(* Logix 5000 project; controller FV vendor 1 type 14 code 217 rev 31.11; software revision 31.00; part 21 of 63 *)
(* tags used below, declared in another part *)
   CheckTimeMask : INT;
   Delphi_Does_Eng_Func : BOOL;
   FR_FV28_AV01 : PlantItem;   // FV28_AV01
   FR_FV28_AV04 : PlantItem;   // FV28_AV04
   FR_FV28_AV05 : PlantItem;   // FV28_AV05
   FR_FV28_AV06 : PlantItem;   // FV28_AV06
   FR_FV28_AV07 : PlantItem;   // FV28_AV07
   FR_FV29_AV01 : PlantItem;   // FV29_AV01
   FR_FV29_AV04 : PlantItem;   // FV29_AV04
   FR_N255 : INT[265];   // CHECKWORDS
   FR_VB1_AV04 : PlantItem;   // VB1_AV04
   FR_VB1_AV05 : PlantItem;   // VB1_AV05
   FR_VB1_AV06 : PlantItem;   // VB1_AV06
   FR_VB1_AV07 : PlantItem;   // VB1_AV07
   FR_VB1_AV08 : PlantItem;   // VB1_AV08
   FR_VB1_AV09 : PlantItem;   // VB1_AV09
   TempChecktime : DINT;
(* FR_Common, continued *)

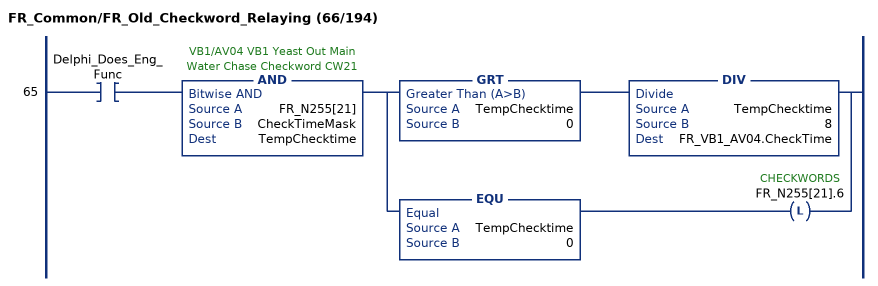
   [picture p370: FR_Common/FR_Old_Checkword_Relaying rungs 65-65]
   65: XIC(Delphi_Does_Eng_Func)AND(FR_N255[21],CheckTimeMask,TempChecktime)[GRT(TempChecktime,0) DIV(TempChecktime,8,FR_VB1_AV04.CheckTime) ,EQU(TempChecktime,0) OTL(FR_N255[21].6) ];
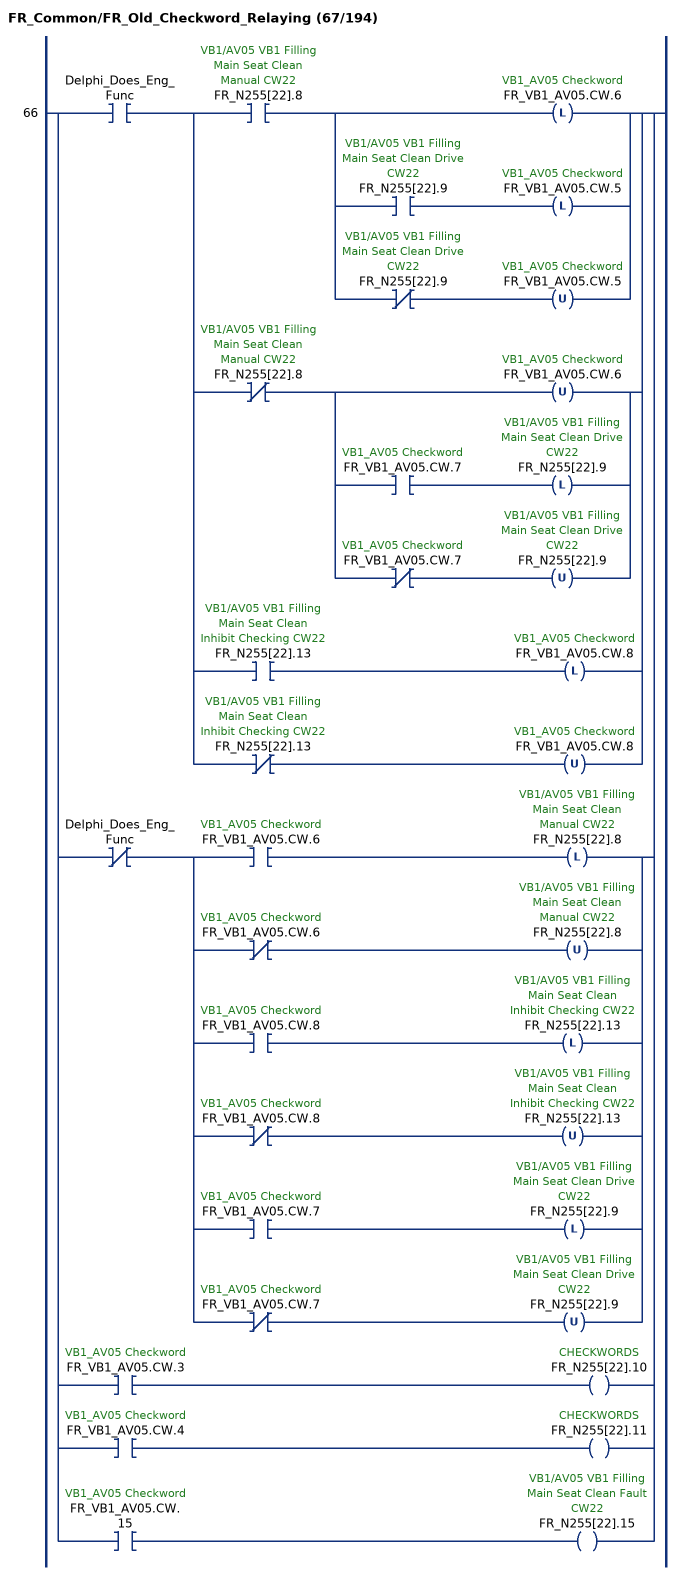
   66: [XIC(Delphi_Does_Eng_Func) [[XIC(FR_N255[22].8) [OTL(FR_VB1_AV05.CW.6) ,XIC(FR_N255[22].9) OTL(FR_VB1_AV05.CW.5) ,XIO(FR_N255[22].9) OTU(FR_VB1_AV05.CW.5) ] ,XIO(FR_N255[22].8) [OTU(FR_VB1_AV05.CW.6) ,[XIC(FR_VB1_AV05.CW.7) OTL(FR_N255[22].9) ,XIO(FR_VB1_AV05.CW.7) OTU(FR_N255[22].9) ] ] ] ,[XIC(FR_N255[22].13) OTL(FR_VB1_AV05.CW.8) ,XIO(FR_N255[22].13) OTU(FR_VB1_AV05.CW.8) ] ] ,XIO(Delphi_Does_Eng_Func) [[XIC(FR_VB1_AV05.CW.6) OTL(FR_N255[22].8) ,XIO(FR_VB1_AV05.CW.6) OTU(FR_N255[22].8) ] ,[XIC(FR_VB1_AV05.CW.8) OTL(FR_N255[22].13) ,XIO(FR_VB1_AV05.CW.8) OTU(FR_N255[22].13) ] ,[XIC(FR_VB1_AV05.CW.7) OTL(FR_N255[22].9) ,XIO(FR_VB1_AV05.CW.7) OTU(FR_N255[22].9) ] ] ,XIC(FR_VB1_AV05.CW.3) OTE(FR_N255[22].10) ,XIC(FR_VB1_AV05.CW.4) OTE(FR_N255[22].11) ,XIC(FR_VB1_AV05.CW.15) OTE(FR_N255[22].15) ];
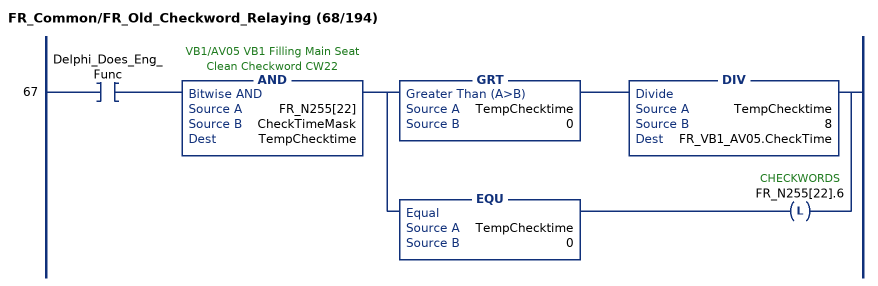
   67: XIC(Delphi_Does_Eng_Func)AND(FR_N255[22],CheckTimeMask,TempChecktime)[GRT(TempChecktime,0) DIV(TempChecktime,8,FR_VB1_AV05.CheckTime) ,EQU(TempChecktime,0) OTL(FR_N255[22].6) ];
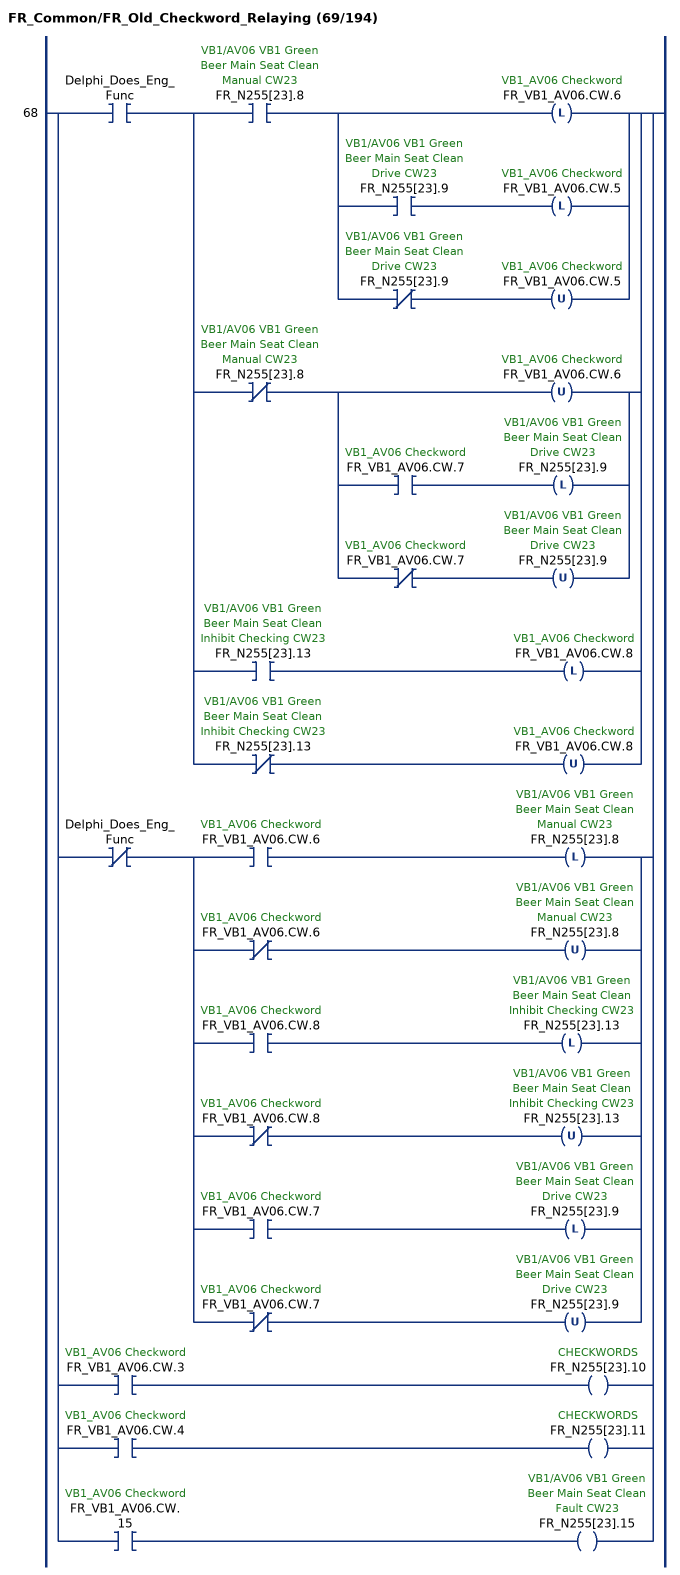
   68: [XIC(Delphi_Does_Eng_Func) [[XIC(FR_N255[23].8) [OTL(FR_VB1_AV06.CW.6) ,XIC(FR_N255[23].9) OTL(FR_VB1_AV06.CW.5) ,XIO(FR_N255[23].9) OTU(FR_VB1_AV06.CW.5) ] ,XIO(FR_N255[23].8) [OTU(FR_VB1_AV06.CW.6) ,[XIC(FR_VB1_AV06.CW.7) OTL(FR_N255[23].9) ,XIO(FR_VB1_AV06.CW.7) OTU(FR_N255[23].9) ] ] ] ,[XIC(FR_N255[23].13) OTL(FR_VB1_AV06.CW.8) ,XIO(FR_N255[23].13) OTU(FR_VB1_AV06.CW.8) ] ] ,XIO(Delphi_Does_Eng_Func) [[XIC(FR_VB1_AV06.CW.6) OTL(FR_N255[23].8) ,XIO(FR_VB1_AV06.CW.6) OTU(FR_N255[23].8) ] ,[XIC(FR_VB1_AV06.CW.8) OTL(FR_N255[23].13) ,XIO(FR_VB1_AV06.CW.8) OTU(FR_N255[23].13) ] ,[XIC(FR_VB1_AV06.CW.7) OTL(FR_N255[23].9) ,XIO(FR_VB1_AV06.CW.7) OTU(FR_N255[23].9) ] ] ,XIC(FR_VB1_AV06.CW.3) OTE(FR_N255[23].10) ,XIC(FR_VB1_AV06.CW.4) OTE(FR_N255[23].11) ,XIC(FR_VB1_AV06.CW.15) OTE(FR_N255[23].15) ];
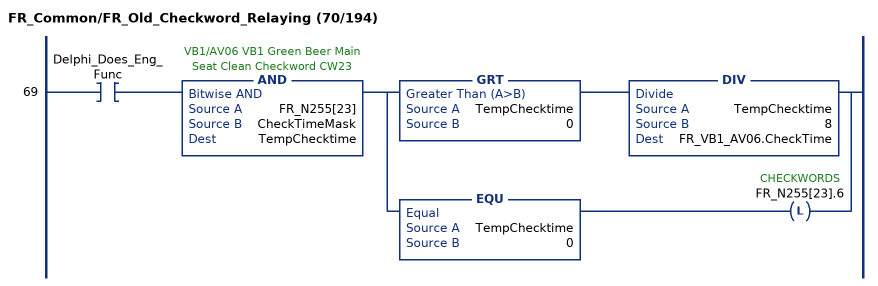
   69: XIC(Delphi_Does_Eng_Func)AND(FR_N255[23],CheckTimeMask,TempChecktime)[GRT(TempChecktime,0) DIV(TempChecktime,8,FR_VB1_AV06.CheckTime) ,EQU(TempChecktime,0) OTL(FR_N255[23].6) ];
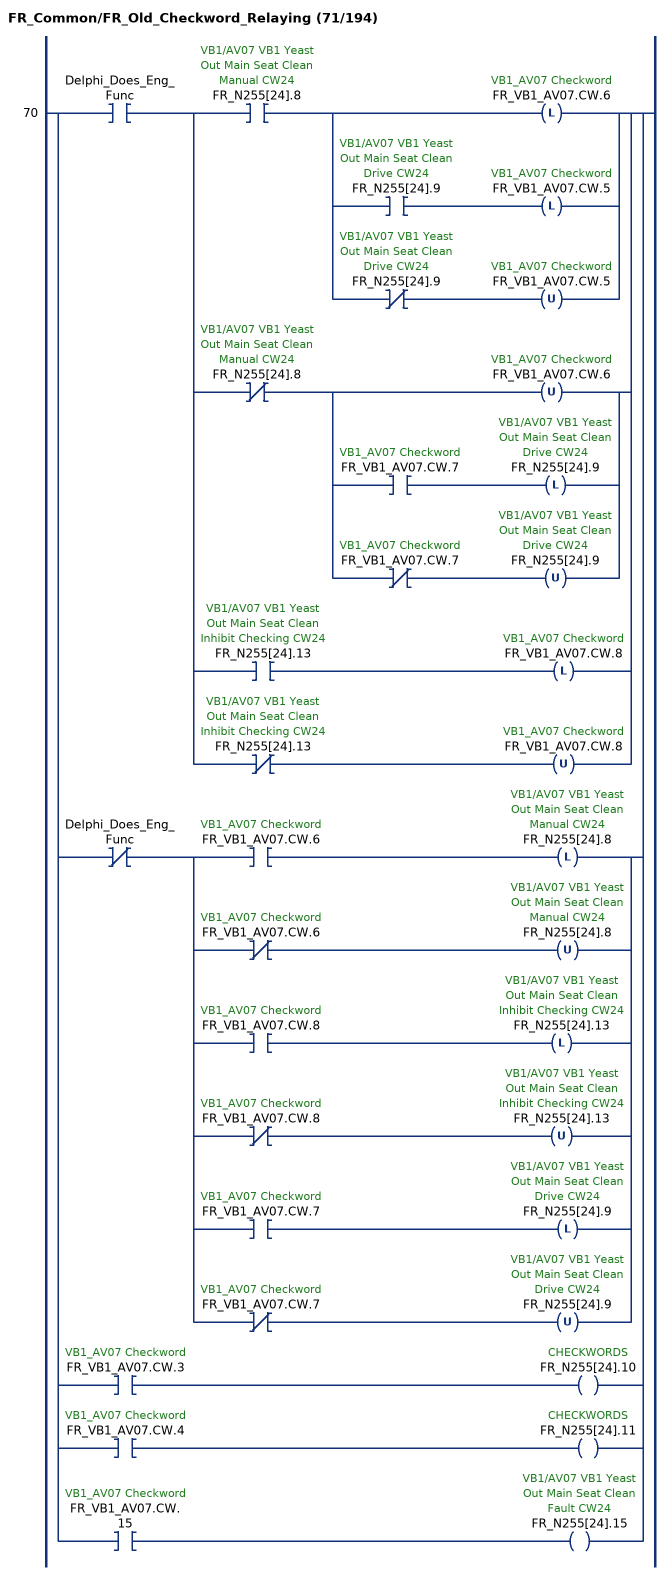
   70: [XIC(Delphi_Does_Eng_Func) [[XIC(FR_N255[24].8) [OTL(FR_VB1_AV07.CW.6) ,XIC(FR_N255[24].9) OTL(FR_VB1_AV07.CW.5) ,XIO(FR_N255[24].9) OTU(FR_VB1_AV07.CW.5) ] ,XIO(FR_N255[24].8) [OTU(FR_VB1_AV07.CW.6) ,[XIC(FR_VB1_AV07.CW.7) OTL(FR_N255[24].9) ,XIO(FR_VB1_AV07.CW.7) OTU(FR_N255[24].9) ] ] ] ,[XIC(FR_N255[24].13) OTL(FR_VB1_AV07.CW.8) ,XIO(FR_N255[24].13) OTU(FR_VB1_AV07.CW.8) ] ] ,XIO(Delphi_Does_Eng_Func) [[XIC(FR_VB1_AV07.CW.6) OTL(FR_N255[24].8) ,XIO(FR_VB1_AV07.CW.6) OTU(FR_N255[24].8) ] ,[XIC(FR_VB1_AV07.CW.8) OTL(FR_N255[24].13) ,XIO(FR_VB1_AV07.CW.8) OTU(FR_N255[24].13) ] ,[XIC(FR_VB1_AV07.CW.7) OTL(FR_N255[24].9) ,XIO(FR_VB1_AV07.CW.7) OTU(FR_N255[24].9) ] ] ,XIC(FR_VB1_AV07.CW.3) OTE(FR_N255[24].10) ,XIC(FR_VB1_AV07.CW.4) OTE(FR_N255[24].11) ,XIC(FR_VB1_AV07.CW.15) OTE(FR_N255[24].15) ];
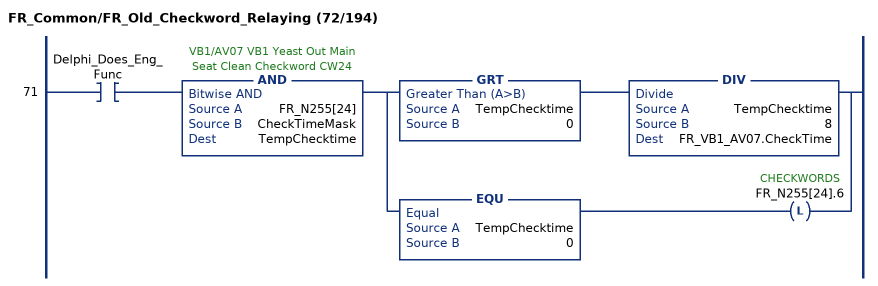
   71: XIC(Delphi_Does_Eng_Func)AND(FR_N255[24],CheckTimeMask,TempChecktime)[GRT(TempChecktime,0) DIV(TempChecktime,8,FR_VB1_AV07.CheckTime) ,EQU(TempChecktime,0) OTL(FR_N255[24].6) ];
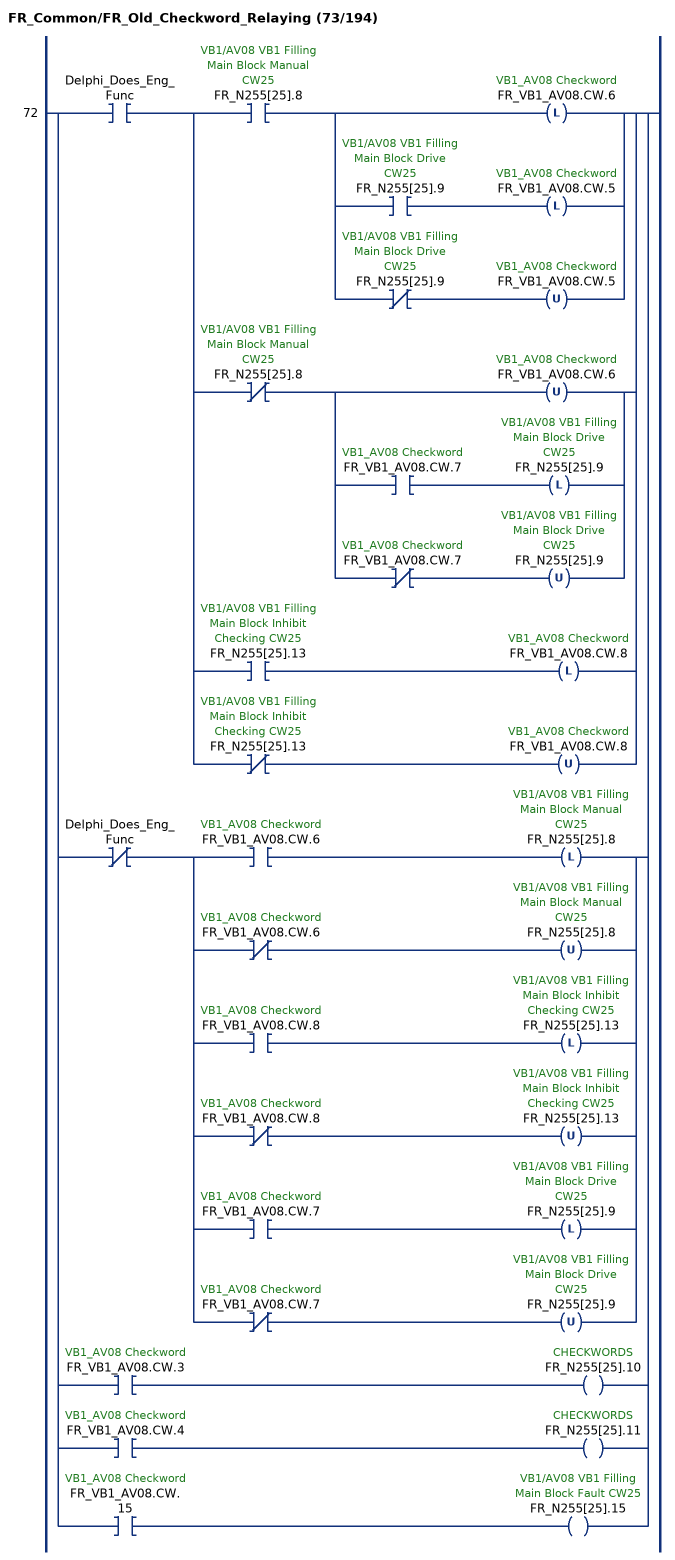
   72: [XIC(Delphi_Does_Eng_Func) [[XIC(FR_N255[25].8) [OTL(FR_VB1_AV08.CW.6) ,XIC(FR_N255[25].9) OTL(FR_VB1_AV08.CW.5) ,XIO(FR_N255[25].9) OTU(FR_VB1_AV08.CW.5) ] ,XIO(FR_N255[25].8) [OTU(FR_VB1_AV08.CW.6) ,[XIC(FR_VB1_AV08.CW.7) OTL(FR_N255[25].9) ,XIO(FR_VB1_AV08.CW.7) OTU(FR_N255[25].9) ] ] ] ,[XIC(FR_N255[25].13) OTL(FR_VB1_AV08.CW.8) ,XIO(FR_N255[25].13) OTU(FR_VB1_AV08.CW.8) ] ] ,XIO(Delphi_Does_Eng_Func) [[XIC(FR_VB1_AV08.CW.6) OTL(FR_N255[25].8) ,XIO(FR_VB1_AV08.CW.6) OTU(FR_N255[25].8) ] ,[XIC(FR_VB1_AV08.CW.8) OTL(FR_N255[25].13) ,XIO(FR_VB1_AV08.CW.8) OTU(FR_N255[25].13) ] ,[XIC(FR_VB1_AV08.CW.7) OTL(FR_N255[25].9) ,XIO(FR_VB1_AV08.CW.7) OTU(FR_N255[25].9) ] ] ,XIC(FR_VB1_AV08.CW.3) OTE(FR_N255[25].10) ,XIC(FR_VB1_AV08.CW.4) OTE(FR_N255[25].11) ,XIC(FR_VB1_AV08.CW.15) OTE(FR_N255[25].15) ];
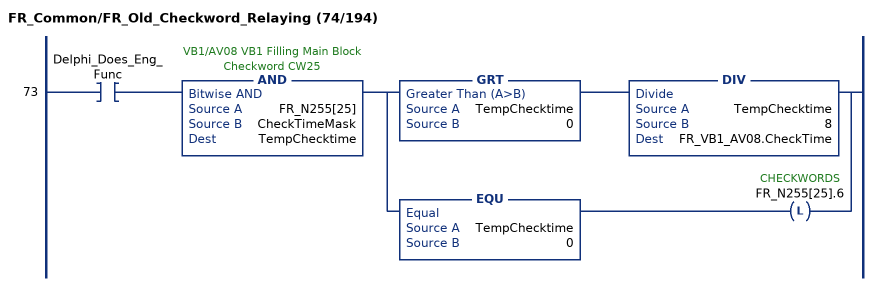
   73: XIC(Delphi_Does_Eng_Func)AND(FR_N255[25],CheckTimeMask,TempChecktime)[GRT(TempChecktime,0) DIV(TempChecktime,8,FR_VB1_AV08.CheckTime) ,EQU(TempChecktime,0) OTL(FR_N255[25].6) ];
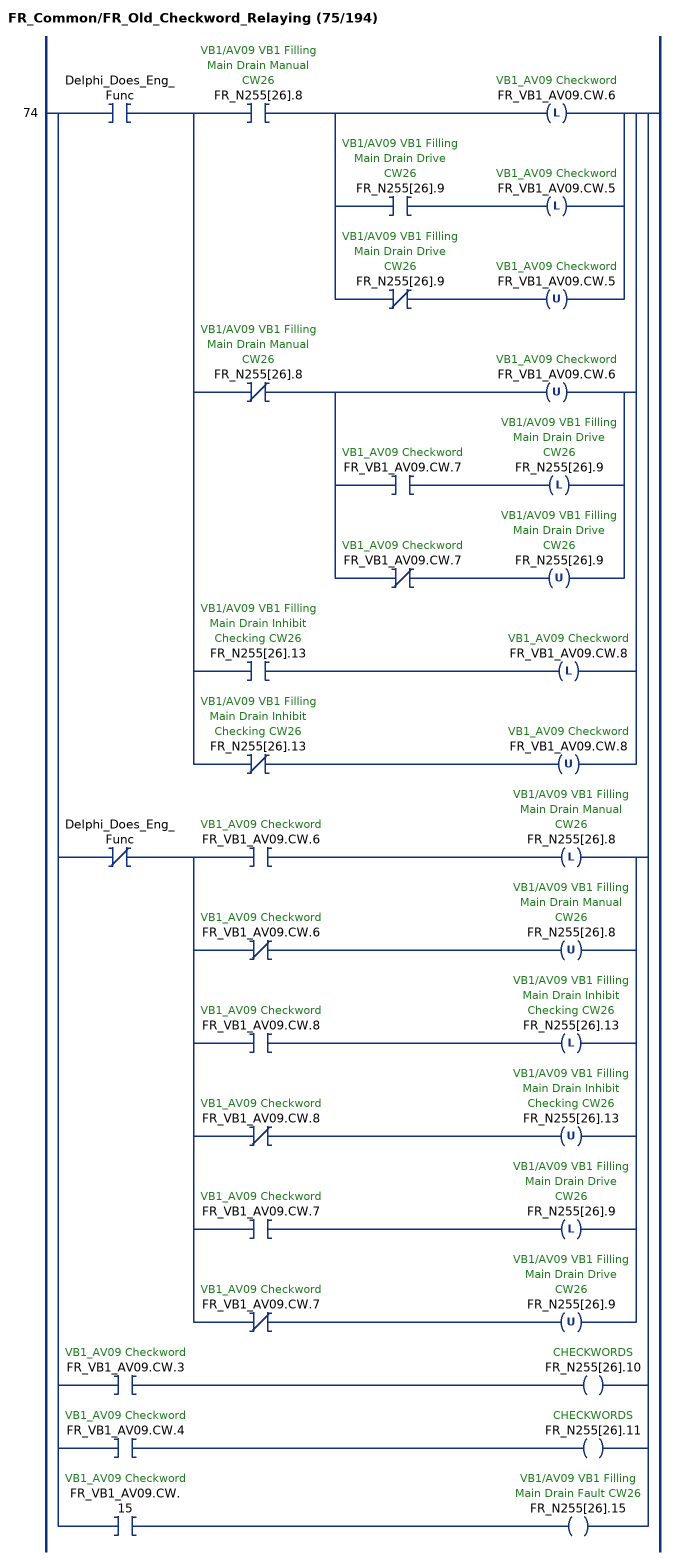
   74: [XIC(Delphi_Does_Eng_Func) [[XIC(FR_N255[26].8) [OTL(FR_VB1_AV09.CW.6) ,XIC(FR_N255[26].9) OTL(FR_VB1_AV09.CW.5) ,XIO(FR_N255[26].9) OTU(FR_VB1_AV09.CW.5) ] ,XIO(FR_N255[26].8) [OTU(FR_VB1_AV09.CW.6) ,[XIC(FR_VB1_AV09.CW.7) OTL(FR_N255[26].9) ,XIO(FR_VB1_AV09.CW.7) OTU(FR_N255[26].9) ] ] ] ,[XIC(FR_N255[26].13) OTL(FR_VB1_AV09.CW.8) ,XIO(FR_N255[26].13) OTU(FR_VB1_AV09.CW.8) ] ] ,XIO(Delphi_Does_Eng_Func) [[XIC(FR_VB1_AV09.CW.6) OTL(FR_N255[26].8) ,XIO(FR_VB1_AV09.CW.6) OTU(FR_N255[26].8) ] ,[XIC(FR_VB1_AV09.CW.8) OTL(FR_N255[26].13) ,XIO(FR_VB1_AV09.CW.8) OTU(FR_N255[26].13) ] ,[XIC(FR_VB1_AV09.CW.7) OTL(FR_N255[26].9) ,XIO(FR_VB1_AV09.CW.7) OTU(FR_N255[26].9) ] ] ,XIC(FR_VB1_AV09.CW.3) OTE(FR_N255[26].10) ,XIC(FR_VB1_AV09.CW.4) OTE(FR_N255[26].11) ,XIC(FR_VB1_AV09.CW.15) OTE(FR_N255[26].15) ];
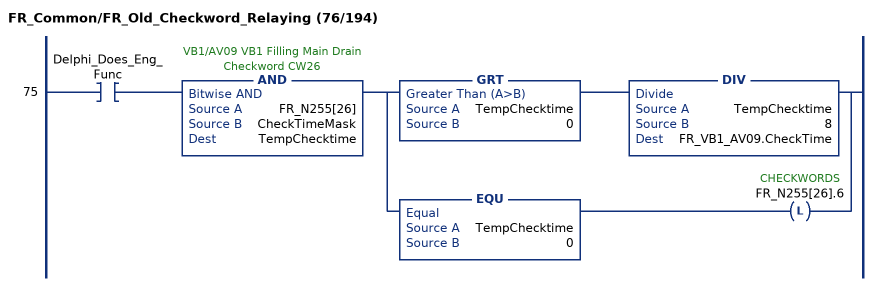
   75: XIC(Delphi_Does_Eng_Func)AND(FR_N255[26],CheckTimeMask,TempChecktime)[GRT(TempChecktime,0) DIV(TempChecktime,8,FR_VB1_AV09.CheckTime) ,EQU(TempChecktime,0) OTL(FR_N255[26].6) ];
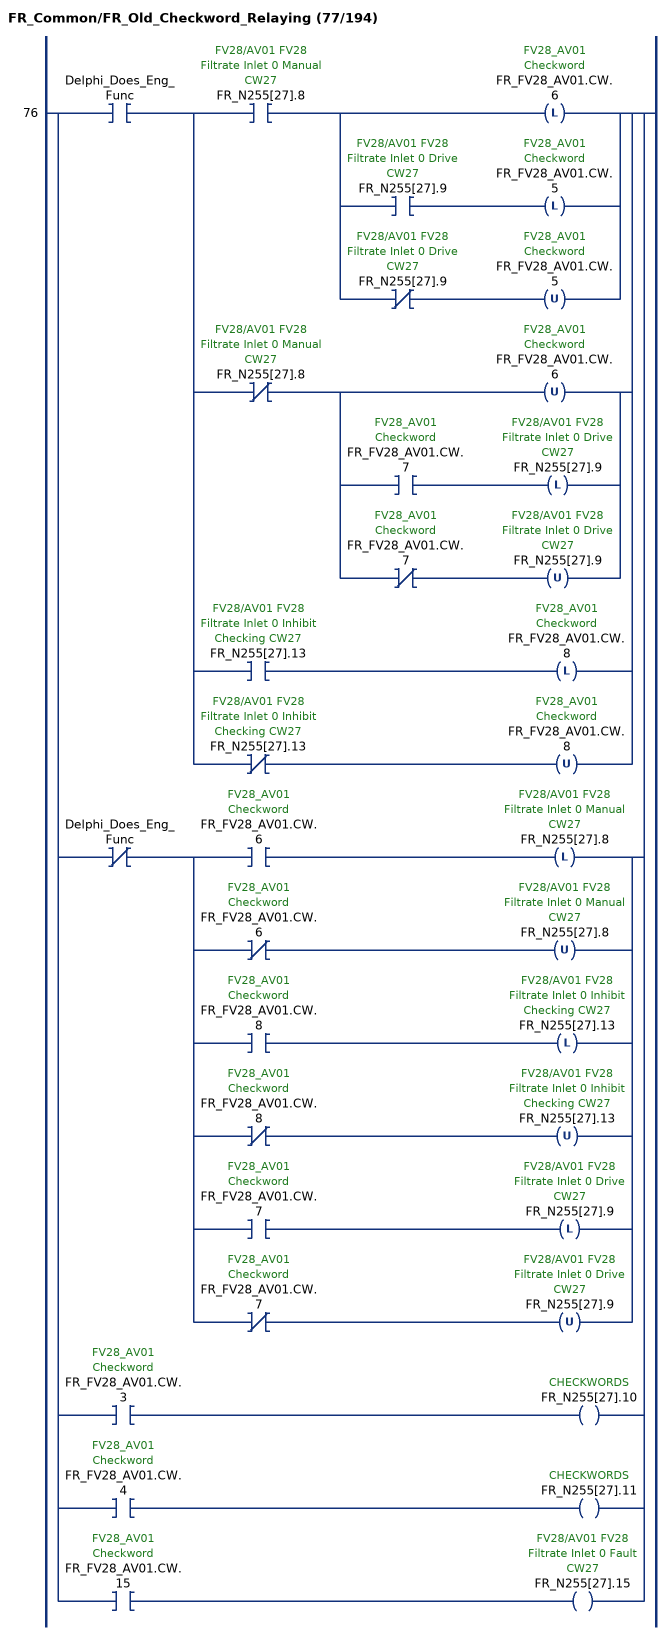
   76: [XIC(Delphi_Does_Eng_Func) [[XIC(FR_N255[27].8) [OTL(FR_FV28_AV01.CW.6) ,XIC(FR_N255[27].9) OTL(FR_FV28_AV01.CW.5) ,XIO(FR_N255[27].9) OTU(FR_FV28_AV01.CW.5) ] ,XIO(FR_N255[27].8) [OTU(FR_FV28_AV01.CW.6) ,[XIC(FR_FV28_AV01.CW.7) OTL(FR_N255[27].9) ,XIO(FR_FV28_AV01.CW.7) OTU(FR_N255[27].9) ] ] ] ,[XIC(FR_N255[27].13) OTL(FR_FV28_AV01.CW.8) ,XIO(FR_N255[27].13) OTU(FR_FV28_AV01.CW.8) ] ] ,XIO(Delphi_Does_Eng_Func) [[XIC(FR_FV28_AV01.CW.6) OTL(FR_N255[27].8) ,XIO(FR_FV28_AV01.CW.6) OTU(FR_N255[27].8) ] ,[XIC(FR_FV28_AV01.CW.8) OTL(FR_N255[27].13) ,XIO(FR_FV28_AV01.CW.8) OTU(FR_N255[27].13) ] ,[XIC(FR_FV28_AV01.CW.7) OTL(FR_N255[27].9) ,XIO(FR_FV28_AV01.CW.7) OTU(FR_N255[27].9) ] ] ,XIC(FR_FV28_AV01.CW.3) OTE(FR_N255[27].10) ,XIC(FR_FV28_AV01.CW.4) OTE(FR_N255[27].11) ,XIC(FR_FV28_AV01.CW.15) OTE(FR_N255[27].15) ];